// TIA Portal project "TESTV18" (V18) (continued)
REGION Network 13: Bit X12 = Allarme 13
   #_w1 := #IV_CND_ALLX12 AND NOT #VW_Allarms.%X12;
   #TI_T12.TON(IN := #_w1, PT := T#5S);
   IF #_w1 AND #TI_T12.Q THEN
       #VW_Allarms.%X12 := TRUE;   // SR flip-flop
   END_IF;
   IF #IV_RST_ALL THEN #VW_Allarms.%X12 := FALSE; END_IF;
END_REGION

REGION Network 14: Bit X13 = Allarme 14
   #_w1 := #IV_CND_ALLX13 AND NOT #VW_Allarms.%X13;
   #TI_T13.TON(IN := #_w1, PT := T#5S);
   IF #_w1 AND #TI_T13.Q THEN
       #VW_Allarms.%X13 := TRUE;   // SR flip-flop
   END_IF;
   IF #IV_RST_ALL THEN #VW_Allarms.%X13 := FALSE; END_IF;
END_REGION

REGION Network 15: Bit X14 = Allarme 15
   #_w1 := #IV_CND_ALLX14 AND NOT #VW_Allarms.%X14;
   #TI_T14.TON(IN := #_w1, PT := T#5S);
   IF #_w1 AND #TI_T14.Q THEN
       #VW_Allarms.%X14 := TRUE;   // SR flip-flop
   END_IF;
   IF #IV_RST_ALL THEN #VW_Allarms.%X14 := FALSE; END_IF;
END_REGION

REGION Network 16: Bit X15 = Allarme 16
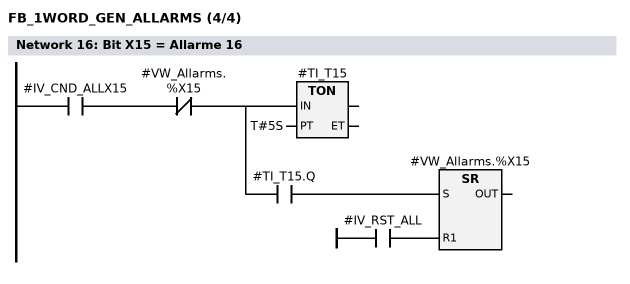
   #_w1 := #IV_CND_ALLX15 AND NOT #VW_Allarms.%X15;
   #TI_T15.TON(IN := #_w1, PT := T#5S);
   IF #_w1 AND #TI_T15.Q THEN
       #VW_Allarms.%X15 := TRUE;   // SR flip-flop
   END_IF;
   IF #IV_RST_ALL THEN #VW_Allarms.%X15 := FALSE; END_IF;
END_REGION
END_FUNCTION_BLOCK

FUNCTION_BLOCK "FB_CYL_DIAGN"   // FB550, LAD
TITLE = FB_CYL_DIAGN
{ S7_Optimized_Access := 'TRUE' }
AUTHOR : C.M.
VERSION : 0.1
// FB per diagnostica cilindro
   VAR_INPUT
      PMI_Limit_Switch_Backward : Bool := FALSE;   // Sensore di posizione cilindro retratto
      PMS_Limit_Switch_Forward : Bool := FALSE;   // Sensore di posizione cilindro esteso
      PST_Home_Position_Backward : Bool := FALSE;   // Posizione HOME indietro
      PST_Home_Position_Forward : Bool := FALSE;   // Posizione HOME avanti
      PST_Latch_In_Backward_Position : Bool := FALSE;   // Interlock in posizione indietro
      PST_Latch_In_Forward_Position : Bool := FALSE;   // Interlock in posizione avanti
      PST_Alarm_Muting : Bool;   // Interlock per sospensione allarmi
      IV_CMD_EV_BCK : Bool;   // Ingresso per conferma attivazione comando cilindro retratto
      IV_CMD_EV_FWD : Bool;   // Ingresso per conferma attivazione comando cilindro esteso
      Station_Info : "Machine_Status_Data";   // Informazioni generali stazione
   END_VAR
   VAR_OUTPUT
      VW_AllarmDIA : Word;   // Variabile WORD per allarmi
   END_VAR
   VAR
      CIN_Auto_Request_Backward : Bool := FALSE;
      CIN_Auto_Request_Forward : Bool := FALSE;
      CIN_Manual_PB_Request_Backward : Bool := FALSE;
      CIN_Manual_PB_Request_Forward : Bool := FALSE;
      CYL_In_Backward_Position : Bool := FALSE;
      CYL_In_Forward_Position : Bool := FALSE;
      CYL_In_Home_Position : Bool := FALSE;
      LOC_SensorBackup_Backward : Bool := FALSE;
      LOC_SensorBackup_Forward : Bool := FALSE;
      LOC_Pulse_1 : Bool;
      LOC_Pulse_2 : Bool;
   END_VAR
   VAR RETAIN
      LOC_DiagnDelay_Backward : Time := T#5s;
      LOC_DiagnDelay_Forward : Time := T#5s;
   END_VAR
   VAR
      LOC_Timer_NotReached_Backward : IEC_TIMER;
      LOC_Timer_NotReached_Forward : IEC_TIMER;
      LOC_Timer_SwitchesContemp : IEC_TIMER;
   END_VAR
   VAR RETAIN
      DIA : "Cylinder_Diagnostic";
   END_VAR
   VAR_TEMP
      No_error : Bool;
   END_VAR
   VAR_TEMP   // added for the SCL form of the ladder/FBD networks
      _w1 : Bool;
   END_VAR
BEGIN

REGION Network 1: *** STATO FINECORSA ***
END_REGION

REGION Network 2: LOGICA - movimento indietro eseguito
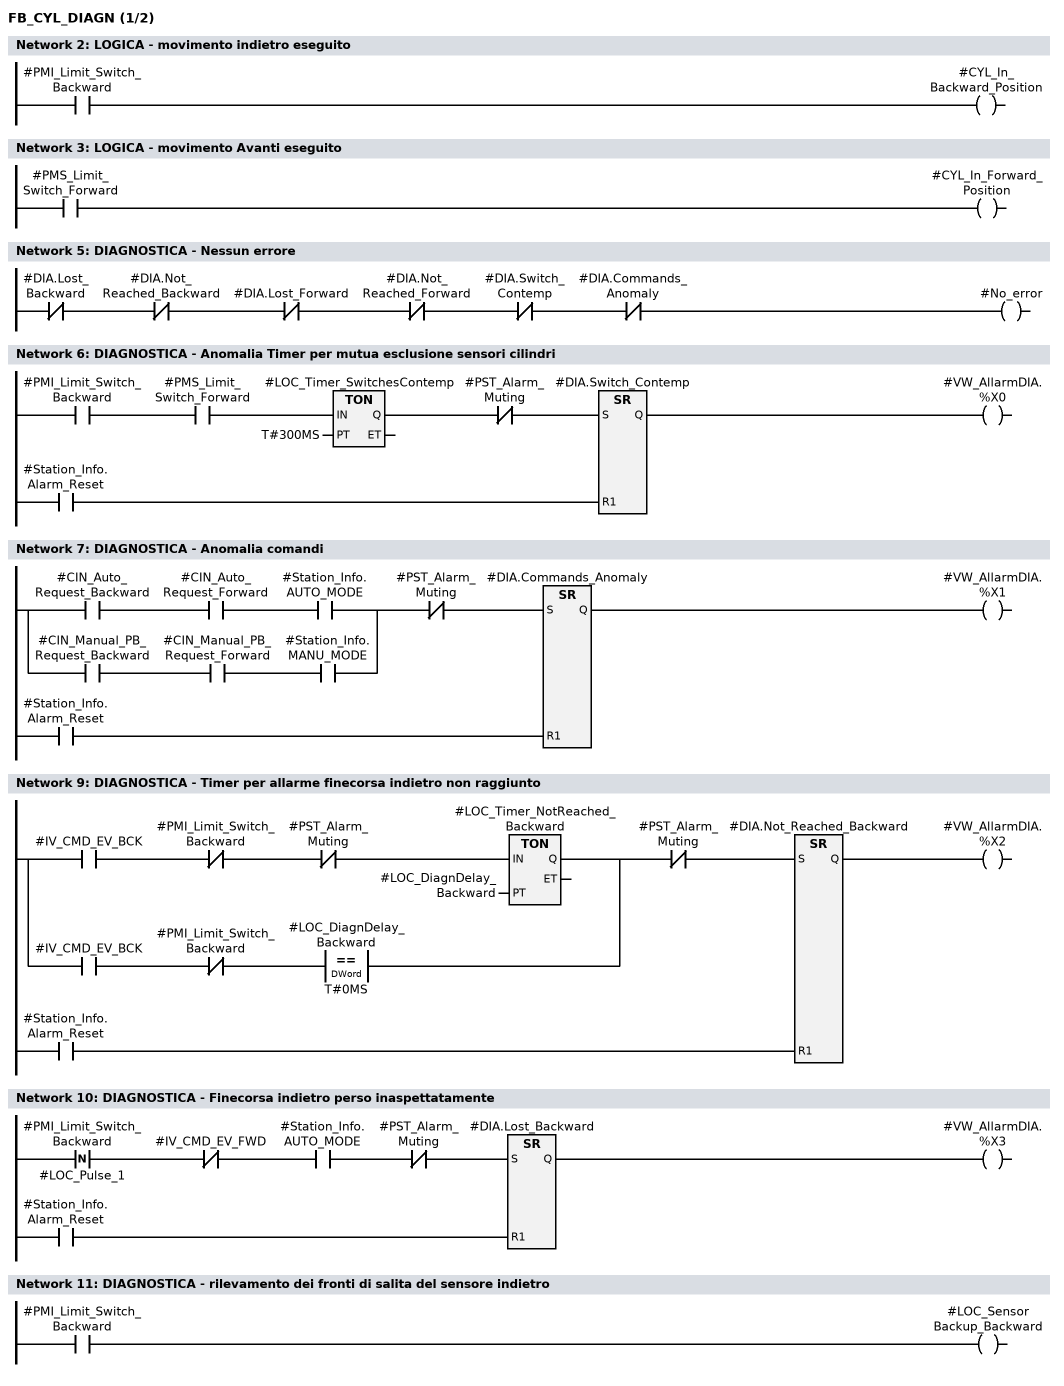
   RUNG wire#powerrail
      Contact( #PMI_Limit_Switch_Backward )
      Coil( #CYL_In_Backward_Position )
   END_RUNG
   // the same network as SCL:
   #CYL_In_Backward_Position := #PMI_Limit_Switch_Backward;
END_REGION

REGION Network 3: LOGICA - movimento Avanti eseguito
   RUNG wire#powerrail
      Contact( #PMS_Limit_Switch_Forward )
      Coil( #CYL_In_Forward_Position )
   END_RUNG
   // the same network as SCL:
   #CYL_In_Forward_Position := #PMS_Limit_Switch_Forward;
END_REGION

REGION Network 4: *** DIAGNOSTICA ***
END_REGION

REGION Network 5: DIAGNOSTICA - Nessun errore
   RUNG wire#powerrail
      I_Contact( #DIA.Lost_Backward )
      I_Contact( #DIA.Not_Reached_Backward )
      I_Contact( #DIA.Lost_Forward )
      I_Contact( #DIA.Not_Reached_Forward )
      I_Contact( #DIA.Switch_Contemp )
      I_Contact( #DIA.Commands_Anomaly )
      Coil( #No_error )
   END_RUNG
   // the same network as SCL:
   #No_error := NOT #DIA.Lost_Backward AND NOT #DIA.Not_Reached_Backward AND NOT #DIA.Lost_Forward AND NOT #DIA.Not_Reached_Forward AND NOT #DIA.Switch_Contemp AND NOT #DIA.Commands_Anomaly;
END_REGION

REGION Network 6: DIAGNOSTICA - Anomalia Timer per mutua esclusione sensori cilindri
   #LOC_Timer_SwitchesContemp.TON(IN := #PMI_Limit_Switch_Backward AND #PMS_Limit_Switch_Forward, PT := T#300MS);
   IF #LOC_Timer_SwitchesContemp.Q AND NOT #PST_Alarm_Muting THEN
       #DIA.Switch_Contemp := TRUE;   // SR flip-flop
   END_IF;
   IF #Station_Info.Alarm_Reset THEN #DIA.Switch_Contemp := FALSE; END_IF;
   #VW_AllarmDIA.%X0 := #DIA.Switch_Contemp;
END_REGION

REGION Network 7: DIAGNOSTICA - Anomalia comandi
   RUNG wire#powerrail
      Contact( #CIN_Auto_Request_Backward )
      Contact( #CIN_Auto_Request_Forward )
      Contact( #Station_Info.AUTO_MODE )
      wire#w1
      I_Contact( #PST_Alarm_Muting )
      S_SR(operand := #DIA.Commands_Anomaly, r1 := wire#w2)
      Coil( #VW_AllarmDIA.%X1 )
   END_RUNG
   RUNG wire#powerrail
      Contact( #CIN_Manual_PB_Request_Backward )
      Contact( #CIN_Manual_PB_Request_Forward )
      Contact( #Station_Info.MANU_MODE )
   END_RUNG wire#w1
   RUNG wire#powerrail
      Contact( #Station_Info.Alarm_Reset )
   END_RUNG wire#w2
   // the same network as SCL:
   IF ((#CIN_Auto_Request_Backward AND #CIN_Auto_Request_Forward AND #Station_Info.AUTO_MODE) OR (#CIN_Manual_PB_Request_Backward AND #CIN_Manual_PB_Request_Forward AND #Station_Info.MANU_MODE)) AND NOT #PST_Alarm_Muting THEN
       #DIA.Commands_Anomaly := TRUE;   // SR flip-flop
   END_IF;
   IF #Station_Info.Alarm_Reset THEN #DIA.Commands_Anomaly := FALSE; END_IF;
   #VW_AllarmDIA.%X1 := #DIA.Commands_Anomaly;
END_REGION

REGION Network 8: *** DIAGNOSTICA SENSORE INDIETRO PMI ***
END_REGION

REGION Network 9: DIAGNOSTICA - Timer per allarme finecorsa indietro non raggiunto
   #LOC_Timer_NotReached_Backward.TON(IN := #IV_CMD_EV_BCK AND NOT #PMI_Limit_Switch_Backward AND NOT #PST_Alarm_Muting,
                           PT := #LOC_DiagnDelay_Backward);
   IF (#LOC_Timer_NotReached_Backward.Q OR (#IV_CMD_EV_BCK AND NOT #PMI_Limit_Switch_Backward AND (#LOC_DiagnDelay_Backward = T#0MS))) AND NOT #PST_Alarm_Muting THEN
       #DIA.Not_Reached_Backward := TRUE;   // SR flip-flop
   END_IF;
   IF #Station_Info.Alarm_Reset THEN #DIA.Not_Reached_Backward := FALSE; END_IF;
   #VW_AllarmDIA.%X2 := #DIA.Not_Reached_Backward;
END_REGION

REGION Network 10: DIAGNOSTICA - Finecorsa indietro perso inaspettatamente
   RUNG wire#powerrail
      N_Contact(operand := #PMI_Limit_Switch_Backward, bit := #LOC_Pulse_1)
      I_Contact( #IV_CMD_EV_FWD )
      Contact( #Station_Info.AUTO_MODE )
      I_Contact( #PST_Alarm_Muting )
      S_SR(operand := #DIA.Lost_Backward, r1 := wire#w1)
      Coil( #VW_AllarmDIA.%X3 )
   END_RUNG
   RUNG wire#powerrail
      Contact( #Station_Info.Alarm_Reset )
   END_RUNG wire#w1
   // the same network as SCL:
   #_w1 := NOT #PMI_Limit_Switch_Backward AND #LOC_Pulse_1;   // falling edge of #PMI_Limit_Switch_Backward
   #LOC_Pulse_1 := #PMI_Limit_Switch_Backward;
   IF #_w1 AND NOT #IV_CMD_EV_FWD AND #Station_Info.AUTO_MODE AND NOT #PST_Alarm_Muting THEN
       #DIA.Lost_Backward := TRUE;   // SR flip-flop
   END_IF;
   IF #Station_Info.Alarm_Reset THEN #DIA.Lost_Backward := FALSE; END_IF;
   #VW_AllarmDIA.%X3 := #DIA.Lost_Backward;
END_REGION

REGION Network 11: DIAGNOSTICA - rilevamento dei fronti di salita del sensore indietro
   RUNG wire#powerrail
      Contact( #PMI_Limit_Switch_Backward )
      Coil( #LOC_SensorBackup_Backward )
   END_RUNG
   // the same network as SCL:
   #LOC_SensorBackup_Backward := #PMI_Limit_Switch_Backward;
END_REGION

REGION Network 12: *** DIAGNOSTICA SENSORE AVANTI PMS ***
END_REGION

REGION Network 13: DIAGNOSTICA - Timer per allarme finecorsa avanti non raggiunto
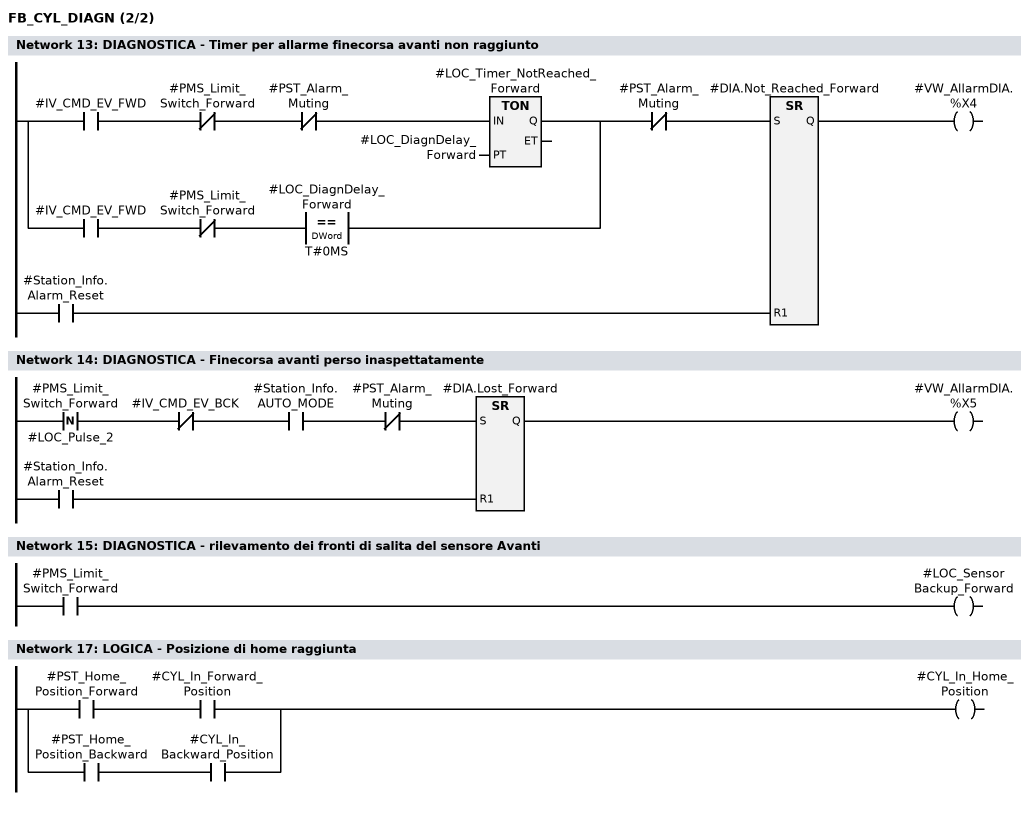
   #LOC_Timer_NotReached_Forward.TON(IN := #IV_CMD_EV_FWD AND NOT #PMS_Limit_Switch_Forward AND NOT #PST_Alarm_Muting,
                           PT := #LOC_DiagnDelay_Forward);
   IF (#LOC_Timer_NotReached_Forward.Q OR (#IV_CMD_EV_FWD AND NOT #PMS_Limit_Switch_Forward AND (#LOC_DiagnDelay_Forward = T#0MS))) AND NOT #PST_Alarm_Muting THEN
       #DIA.Not_Reached_Forward := TRUE;   // SR flip-flop
   END_IF;
   IF #Station_Info.Alarm_Reset THEN #DIA.Not_Reached_Forward := FALSE; END_IF;
   #VW_AllarmDIA.%X4 := #DIA.Not_Reached_Forward;
END_REGION

REGION Network 14: DIAGNOSTICA - Finecorsa avanti perso inaspettatamente
   RUNG wire#powerrail
      N_Contact(operand := #PMS_Limit_Switch_Forward, bit := #LOC_Pulse_2)
      I_Contact( #IV_CMD_EV_BCK )
      Contact( #Station_Info.AUTO_MODE )
      I_Contact( #PST_Alarm_Muting )
      S_SR(operand := #DIA.Lost_Forward, r1 := wire#w1)
      Coil( #VW_AllarmDIA.%X5 )
   END_RUNG
   RUNG wire#powerrail
      Contact( #Station_Info.Alarm_Reset )
   END_RUNG wire#w1
   // the same network as SCL:
   #_w1 := NOT #PMS_Limit_Switch_Forward AND #LOC_Pulse_2;   // falling edge of #PMS_Limit_Switch_Forward
   #LOC_Pulse_2 := #PMS_Limit_Switch_Forward;
   IF #_w1 AND NOT #IV_CMD_EV_BCK AND #Station_Info.AUTO_MODE AND NOT #PST_Alarm_Muting THEN
       #DIA.Lost_Forward := TRUE;   // SR flip-flop
   END_IF;
   IF #Station_Info.Alarm_Reset THEN #DIA.Lost_Forward := FALSE; END_IF;
   #VW_AllarmDIA.%X5 := #DIA.Lost_Forward;
END_REGION

REGION Network 15: DIAGNOSTICA - rilevamento dei fronti di salita del sensore Avanti
   RUNG wire#powerrail
      Contact( #PMS_Limit_Switch_Forward )
      Coil( #LOC_SensorBackup_Forward )
   END_RUNG
   // the same network as SCL:
   #LOC_SensorBackup_Forward := #PMS_Limit_Switch_Forward;
END_REGION

REGION Network 16: *** SEGMENTI DI LOGICA AUSILIARI ***
END_REGION

REGION Network 17: LOGICA - Posizione di home raggiunta
   RUNG wire#powerrail
      Contact( #PST_Home_Position_Forward )
      Contact( #CYL_In_Forward_Position )
      wire#w1
      Coil( #CYL_In_Home_Position )
   END_RUNG
   RUNG wire#powerrail
      Contact( #PST_Home_Position_Backward )
      Contact( #CYL_In_Backward_Position )
   END_RUNG wire#w1
   // the same network as SCL:
   #CYL_In_Home_Position := (#PST_Home_Position_Forward AND #CYL_In_Forward_Position) OR (#PST_Home_Position_Backward AND #CYL_In_Backward_Position);
END_REGION
END_FUNCTION_BLOCK

// folder: LGF/1 Date and timer operations

FUNCTION "LGF_GetCalendarDay" : DInt   // FC10028, SCL
TITLE = LGF_GetCalendarDay
{ S7_Optimized_Access := 'TRUE' }
AUTHOR : Siemens_Digital_Industry
FAMILY : LGF
NAME : LGF_GetCalendarDay
// This function uses the specified date to calculate the number of days that have passed since the beginning of the year (1st January).
// 
// The function is used in the functions “LGF_GetCalendarWeek_ISO” and “LGF_GetCalendarWeek_US”.
// Diese Funktion berechnet aus dem vorgegebenen Datum die Anzahl der Tage, die seit dem Anfang des Jahres vergangen sind (1. Januar).
// 
// Die Funktion wird in den Funktionen "LGF_GetCalendarWeek_ISO" und "LGF_GetCalendarWeek_US" verwendet.
   VAR_INPUT
      "date" : DTL;   // Date for the calculation of the calendar days since 1 January. / Datum für die Berechnung der vergangenen Kalendertagen seit dem 01. Januar
   END_VAR
   VAR_OUTPUT
      error : Bool;   // FALSE: No error / TRUE: An error occurred during the execution of the FB / FALSE: Kein Fehler / TRUE: Während der Ausführung des FB ist ein Fehler aufgetreten
      status : Word;   // 16#0000-16#7FFF: Status of the FB / 16#8000-16#FFFF: Error identification (see following Table) / 16#0000-16#7FFF: Status des FB / 16#8000-16#FFFF: Fehleridentifikation (siehe folgende Tabelle)
   END_VAR
   VAR_TEMP
      tempDaysPassed : DInt;   // Temp tag for the number of days past / Temp Variable für die Anzahl der vergangenen Tage
      tempDate : DTL;   // Temp variable to store date for calculations / Temp Variable um Datum für Berechung zwischen zu speichern
   END_VAR
   // Ret_Val : Days past since January 1st. / Vergangene Tage seit 1. Januar.
   VAR CONSTANT
      FIRST_DAY : USInt := 1;   // 1st of a month / 1. Tag eines Monats
      LAST_DAY : USInt := 31;   // 31st of a month / 31. Tag eines Monats
      JANUARY : USInt := 1;   // Month number for January / Monatsnumer Januar
      DECEMBER : USInt := 12;   // Month number for December / Monatsnummer Dezember
      TIME_ZERO_FORCE_UPDATE : Time := t#0d;   // By adding zero an update of DTL Tag is forced and auto checks are applied / Durch die Addition von "0" wird ein Update üder den Zeitstemple erstellt und ebenfalls auf gültigkeit geprüft.
      ONE_DAY : DInt := 1;   // One single day for incrementing / Ein Tag für inkrementierungen
      STATUS_NO_ERROR : Word := 16#0000;   // Status: no error occurred / Status: kein Fehler aufgetreten
      ERR_LIM_DATE : Word := 16#8201;   // Date out of the range, has to be greater than <1970-01-01 ; 2262-04-11> / Datum ausserhalb des gültigen Bereiches, es muss nach dem <1970-01-01 ; 2262-04-11> liegen
   END_VAR
BEGIN
   REGION BLOCK INFO HEADER
     //===============================================================================
     // SIEMENS AG / (c)Copyright 2019
     //-------------------------------------------------------------------------------
     // Title:            LGF_GetCalendarDay
     // Comment/Function: This function calculates for a date the passed days since 1st January.
     // Library/Family:   LGF(Library General Functions)
     // Author:           Siemens Digital Industry Support
     // Tested with:      S7-PLCSIM Advanced V2.0 SP1
     // Engineering:      TIA Portal V15.1
     // Restrictions:     ENO disabled - error handling done with error and status
     // Requirements:     PLC (S7-1200 / S7-1500)
     //-------------------------------------------------------------------------------
     // Change log table:
     // Version  | Date       | Expert in charge       | Changes applied
     //----------|------------|------------------------|------------------------------
     // 01.00.00 16.07.2019  Simatic Systems Support
     //                      First release
     //                      ENO used for internal error handling, interface has error and status
     //                      temp tag naming, insert constant
     // 03.00.00 23.04.2020  Simatic Systems Support
     //                      Set version to V3.0.0, harmonize the version of the whole library
     // 03.00.01 19.01.2020  Simatic Systems Support
     //                      Insert documentation
     //=============================================================================
   END_REGION BLOCK INFO HEADER

   REGION INITIALISATION
     #tempDate := #date;
     #tempDaysPassed := 0;
   END_REGION

   REGION COUNT DAYS
     // Check #date
     // adding zero forces the PLC to update the tag and eno check
     #tempDate := #tempDate + #TIME_ZERO_FORCE_UPDATE;
     IF ENO = FALSE THEN
       #error := TRUE;
       #status := #ERR_LIM_DATE;
       #LGF_GetCalendarDay := #tempDaysPassed;
       RETURN;
     END_IF;

     // Weekday of 1st January in the current year
     #tempDate.MONTH := #JANUARY;
     #tempDate.DAY := #FIRST_DAY;
     // adding zero forces the PLC to update the tag
     // in this case especially the weekday
     #tempDate := #tempDate + #TIME_ZERO_FORCE_UPDATE;

     // Days passed in the year since 1st January, "date" included
     #tempDaysPassed := DATE_TO_DINT(DTL_TO_DATE(#date)) - DATE_TO_DINT(DTL_TO_DATE(#tempDate)) + #ONE_DAY;
   END_REGION

   REGION OUTPUTS
     #error := FALSE;
     #status := #STATUS_NO_ERROR;
     #LGF_GetCalendarDay := #tempDaysPassed;

     // ENO is not used, forced to TRUE
     ENO := TRUE;
   END_REGION
END_FUNCTION

// folder: LGF/4 Math operations

FUNCTION "LGF_CalcDistance_2D" : LReal   // FC10020, SCL
TITLE = LGF_CalcDistance_2D
{ S7_Optimized_Access := 'TRUE' }
AUTHOR : Siemens_Digital_Industries
FAMILY : LGF
NAME : LGF_CalcDistance_2D
// The function calculates the distance between two points in the plane. / Die Funktion berechnet den Abstand zwischen zwei Punkten in der Ebene.
   VAR_INPUT
      x1 : LReal;   // X coordinate point 1 / X Koordinate Punkt 1
      y1 : LReal;   // Y coordinate point 1 / Y Koordinate Punkt 1
      x2 : LReal;   // X coordinate point 2 / X Koordinate Punkt 2
      y2 : LReal;   // Y coordinate point 2 / Y Koordinate Punkt 2
   END_VAR
   // Ret_Val : Calculated distance between the Points / Berechnete Distanz zwischen den Punkten
BEGIN
   REGION Block info header
     //=============================================================================
     // Siemens AG / (c)Copyright 2017
     //-----------------------------------------------------------------------------
     // Title:            LGF_CalcDistance_2D
     // Comment/Function: Calculates the distance between two points in 2D space
     // Library/Family:   LGF(Library General Functions)
     // Author:           Siemens Digital Industry Support
     // Tested with:      S7-PLCSIM Advanced V2.0 SP1
     // Engineering:      TIA Portal V15 Update 2
     // Restrictions:     ENO disabled - ENO mechanism is not used
     // Requirements:     PLC (S7-1200 / S7-1500)
     //-------------------------------------------------------------------------------
     // Change log table:
     // Version  | Date       | Expert in charge       | Changes applied
     //----------|------------|------------------------|------------------------------
     // 01.00.00 06.07.2018  Siemens Industry Online Support
     //                      First released version
     // 01.00.01 17.08.2018  Siemens Industry Online Support
     //                      Upgrade: TIA V15 Update 2
     // 01.00.02 23.11.2018  Siemens Industry Online Support
     //                      Upgrade: TIA V15.1
     // 01.02.00 04.10.2019  Simatic Systems Support
     //                      renamed from "Distance" to "CalcDistance_2D"
     //                      Data type changed to LREAL
     //                      Data type changed to LREAL
     // 03.00.00 23.04.2020  Simatic Systems Support
     //                      Set version to V3.0.0, harmonize the version of the whole library
     // 03.00.01 12.11.2020  Simatic Systems Support
     //                      Insert documentation
     //=============================================================================
   END_REGION Block info header

   REGION DESCRIPTION
     (/*The block calculates the distance between two points in a Cartesian coordinate system. The distance is calculated with the following formula:

   $$
    result = \sqrt[2]{(x_2-x_1)^2+(y_2-y_1)^2}
   $$

   ------

   Figure: Graphical representation

   ![LGF_CalcDistance_2D - Principle of operation](LGF_CalcDistance_2D.PNG "LGF_CalcDistance_2D - Principle of operation")
   Der Baustein berechnet den Abstand zwischen zwei Punkten in einem kartesischen Koordinatensystem. Der Abstand wird mit nachfolgender Formel berechnet:

   $$
    result = \sqrt[2]{(x_2-x_1)^2+(y_2-y_1)^2}
   $$

   ------

   Abbildung: Graphische Darstellung

   ![LGF_CalcDistance_2D - Funktionsweise](LGF_CalcDistance_2D.PNG "LGF_CalcDistance_2D - Funktionsweise")*/)
   END_REGION DESCRIPTION

   REGION Program
     // Calculating the distance
     #LGF_CalcDistance_2D := SQRT(SQR(#x2 - #x1) + SQR(#y2 - #y1));
     // ENO mechanism is not used
     ENO := TRUE;
   END_REGION
END_FUNCTION

// folder: LGF/6 Converter operations

FUNCTION "LGF_BinaryToGray" : DWord   // FC10021, SCL
TITLE = LGF_BinaryToGray
{ S7_Optimized_Access := 'TRUE' }
AUTHOR : Siemens_Digital_Industry
FAMILY : LGF
NAME : LGF_BinaryToGray
// This function converts a binary coded value into a Gray-coded value. / Diese Funktion wandelt einen binär codierten Wert in einen Gray codierten Wert um.
   VAR_INPUT
      variableBinary : DWord;   // Binary coded value to convert to Gray code / Binär codierter Wert der zu Gray-Code umgerechnet wird
   END_VAR
   // Ret_Val : Gray-coded value / Gray codierter Wert
   VAR CONSTANT
      BIT_SHIFT_1 : USInt := 1;   // The number (1) of bit positions by which the specified value should be shifted.
   END_VAR
BEGIN
   REGION BLOCK INFO HEADER
     //===============================================================================
     // SIEMENS AG / (c)Copyright 2017
     //-------------------------------------------------------------------------------
     // Title:            LGF_BinaryToGray
     // Comment/Function: This function converts a binary value to a gray coded value
     // Library/Family:   LGF(Library General Functions)
     // Author:           Siemens Digital Industry Support
     // Tested with:      CPU1212C DC/DC/DC FW:V4.2
     // Engineering:      TIA Portal V14 Update 1
     // Restrictions:     ENO disabled - no error handling needed
     // Requirements:     PLC (S7-1200 / S7-1500)
     //-------------------------------------------------------------------------------
     // Change log table:
     // Version  | Date       | Expert in charge       | Changes applied
     //----------|------------|------------------------|------------------------------
     // 01.00.00 | 19.08.2015 | Siemens Industry Online Support
     //                         First released version
     // 01.00.01 | 28.10.2015 | Siemens Industry Online Support
     //                         Name changed
     // 01.00.02 | 02.01.2017 | Siemens Industry Online Support
     //                         Upgrade: TIA Portal V14 Update 1
     // 01.00.03 | 17.08.2018 | Siemens Industry Online Support
     //                         Upgrade: TIA V15 Update 2
     // 01.00.04 | 23.11.2018 | Siemens Industry Online Support
     //                         Upgrade: TIA V15.1
     // 01.00.05 | 11.06.2019 | Simatic Systems Support
     //                         Standard header and block parameters update
     //                         Add ENO handling
     // 03.00.00 | 23.04.2020 | Simatic Systems Support | Set version to V3.0.0
     //                         Harmonize the version of the whole library
     // 03.00.01 | 23.02.2021 | Simatic Systems Support
     //                         Insert documentation
     //===============================================================================
   END_REGION Block info header

   REGION OUTPUTS
     #LGF_BinaryToGray := #variableBinary XOR SHR(IN := #variableBinary, N := #BIT_SHIFT_1);

     // no error handling needed
     ENO := TRUE;
   END_REGION
END_FUNCTION

// folder: LGF/6 Converter operations/Binary types - Split/Merge

FUNCTION "LGF_MergeBitsToByte" : Byte   // FC10060, SCL
TITLE = LGF_MergeBitsToByte
{ S7_Optimized_Access := 'TRUE' }
AUTHOR : Siemens_Digital_Industry
FAMILY : LGF
NAME : LGF_MergeBitsToByte
// This function merge 8 Bits / 8 Boolean variables into one Byte variable. / Diese Funktion führt 8 Bit / 8 Boolsche Variablen in einer Byte Variable zusammen.
   VAR_INPUT
      bit7 : Bool;   // Input Bit 7 - MSB
      bit6 : Bool;   // Input Bit 6
      bit5 : Bool;   // Input Bit 5
      bit4 : Bool;   // Input Bit 4
      bit3 : Bool;   // Input Bit 3
      bit2 : Bool;   // Input Bit 2
      bit1 : Bool;   // Input Bit 1
      bit0 : Bool;   // Input Bit 0 - LSB
   END_VAR
   VAR_TEMP
      tempByte : Byte;   // Temp memory to merge Bits into a Byte / Temp speicher zum zusammenführen der Bits zu einem Byte
   END_VAR
   // Ret_Val : Composite Bit sequence stored as Byte variable / Zusammengefügte Bitfolge, gespeichert in einer Byte Variable
BEGIN
   REGION BLOCK INFO HEADER
     //===============================================================================
     // SIEMENS AG / (c)Copyright 2018
     //-------------------------------------------------------------------------------
     // Title:            LGF_MergeBitsToByte
     // Comment/Function: This function merge 8 Bits / 8 Boolean variables into one Byte variable.
     // Library/Family:   LGF (Library General Functions)
     // Author:           Siemens Digital Industry Support
     // Tested with:      S7-PLCSIM Advanced V2.0 SP1
     // Engineering:      TIA Portal V14 / V14SP1
     // Restrictions:     ENO disabled - no error handling, no failure possible.
     // Requirements:     PLC (S7-1200 / S7-1500)
     //-------------------------------------------------------------------------------
     // Change log table:
     // Version  | Date       | Expert in charge       | Changes applied
     //----------|------------|------------------------|------------------------------
     // 01.00.00 | 20.06.2019 | Simatic Systems Support
     //                         First release
     // 03.00.00 | 23.04.2020 | Simatic Systems Support | Set version to V3.0.0
     //                         harmonize the version of the whole library
     // 03.00.01 | 22.02.2021 | Simatic Systems Support
     //                         Insert documentation
     //=============================================================================
   END_REGION

   REGION MERGE
     // set the bits by slice access
     #tempByte.%X7 := #bit7;
     #tempByte.%X6 := #bit6;
     #tempByte.%X5 := #bit5;
     #tempByte.%X4 := #bit4;
     #tempByte.%X3 := #bit3;
     #tempByte.%X2 := #bit2;
     #tempByte.%X1 := #bit1;
     #tempByte.%X0 := #bit0;
   END_REGION

   REGION OUTPUT
     #LGF_MergeBitsToByte := #tempByte;
     // no error handling needed
     ENO := TRUE;
   END_REGION
END_FUNCTION

FUNCTION "LGF_SplitByteToBits" : Void   // FC10063, SCL
TITLE = LGF_SplitByteToBits
{ S7_Optimized_Access := 'TRUE' }
AUTHOR : Siemens_Digital_Industry
FAMILY : LGF
NAME : LGF_SplitByteToBits
// This function splits a Byte variable into 8 Boolean / 8 Bit variables. / Diese Funktion zerlegt eine Byte Variable in 8 Bool / 8 Bit Variablen.
   VAR_INPUT
      "byte" : Byte;   // Bit sequence to be split / Bitfolge die zerlegt wird
   END_VAR
   VAR_OUTPUT
      bit7 : Bool;   // Output Bit 7 - MSB
      bit6 : Bool;   // Output Bit 6
      bit5 : Bool;   // Output Bit 5
      bit4 : Bool;   // Output Bit 4
      bit3 : Bool;   // Output Bit 3
      bit2 : Bool;   // Output Bit 2
      bit1 : Bool;   // Output Bit 1
      bit0 : Bool;   // Output Bit 0 - LSB
   END_VAR
BEGIN
   REGION BLOCK INFO HEADER
     //===============================================================================
     // SIEMENS AG / (c)Copyright 2018
     //-------------------------------------------------------------------------------
     // Title:            LGF_SplitByteToBits
     // Comment/Function: This function splits a Byte variable into 8 Boolean / 8 Bit variables
     // Library/Family:   LGF (Library General Functions)
     // Author:           Siemens Digital Industry Support
     // Tested with:      S7-PLCSIM Advanced V2.0 SP1
     // Engineering:      TIA Portal V14 / V14SP1
     // Restrictions:     ENO disabled - no error handling, no failure possible.
     // Requirements:     PLC (S7-1200 / S7-1500)
     //-------------------------------------------------------------------------------
     // Change log table:
     // Version  | Date       | Expert in charge       | Changes applied
     //----------|------------|------------------------|------------------------------
     // 01.00.00 | 20.06.2019 | Simatic Systems Support
     //                         First release
     // 03.00.00 | 23.04.2020 | Simatic Systems Support | Set version to V3.0.0
     //                         harmonize the version of the whole library
     // 03.00.01 | 22.02.2021 | Simatic Systems Support
     //                         Insert documentation
     //=============================================================================
   END_REGION

   REGION OUTPUT
     // get the bits by slice access
     #bit7 := #byte.%X7;
     #bit6 := #byte.%X6;
     #bit5 := #byte.%X5;
     #bit4 := #byte.%X4;
     #bit3 := #byte.%X3;
     #bit2 := #byte.%X2;
     #bit1 := #byte.%X1;
     #bit0 := #byte.%X0;
     // no error handling needed
     ENO := TRUE;
   END_REGION
END_FUNCTION

// folder: MTA/Vari

FUNCTION_BLOCK "ALM_VALVE_CFG1"   // FB2, LAD
TITLE = FB gestione allarmi elettrov. con cilindro pneum.
{ S7_Optimized_Access := 'TRUE' }
AUTHOR : Cecini_M
VERSION : 0.1
// ROUTINE DI GESTIONE ALLARMI ELETTROVALVOLA COMBINATA CON CILINDRO PNEUMATICO.
//  - Usare ingressi CMD1 e CMD2 per bistabile. Usare negazione di CMD1 su CMD2 per monost.
//  - Ingressi di timeout in S 0.0 (convertiti all'interno dell'FB)
//  - 2 CMD Valvola + 2 Sensori posizione SM
//  - Allarme mancanza sensore su CMD1
//  - Allarme mancanza sensore su CMD2
//  - Allarme mutua eslusione entrambi SM
   VAR_INPUT
      IV_YV_CMD1 : Bool;   // Ingresso comando direzione 1
      IV_YV_CMD2 : Bool;   // Ingresso comando direzione 2
      IV_FBK_CMD1 : Bool;   // Ingresso sensore SM comando direzione 1
      IV_FBK_CMD2 : Bool;   // Ingresso sensore SM comando direzione 1
   END_VAR
   VAR_OUTPUT
      Vb_ALM1 : Bool;
      Vb_ALM2 : Bool;
      Vb_ALM3 : Bool;
   END_VAR
   VAR_IN_OUT
      IV_ACK_ALM1 : Bool;   // Ingresso ACK riconoscimento ALM1
      IV_ACK_ALM2 : Bool;   // Ingresso ACK riconoscimento ALM2
      IV_ACK_ALM3 : Bool;   // Ingresso ACK riconoscimento ALM3
      TI_ToutALM1 : UInt;   // Timeout allarme1
      TI_ToutALM2 : UInt;   // Timeout allarme2
      TI_ToutALM3 : UInt;   // Timeout allarme3
   END_VAR
   VAR
      TI_T1 : IEC_TIMER;   // Timer ALM1
      TI_T2 : IEC_TIMER;   // Timer ALM1
      TI_T3 : IEC_TIMER;   // Timer ALM1
      ME_ALM1 : Bool;   // Memoria allarme 1 SM CMD1
      ME_ALM2 : Bool;   // Memoria allarme 2 SM CMD2
      ME_ALM3 : Bool;   // Memoria allarme 3 mutua esclusione sensori SM
      VA_SetP_TIALM1 : DInt;   // Valore di SETPOINT per timer ALM1
      VA_SetP_TIALM2 : DInt;   // Valore di SETPOINT per timer ALM2
      VA_SetP_TIALM3 : DInt;   // Valore di SETPOINT per timer ALM3
   END_VAR
   VAR_TEMP
      VA_AppRis1 : UInt;   // Variabile appoggio risultato intermedio 1
      VA_AppRis2 : UInt;   // Variabile appoggio risultato intermedio 2
      VA_AppRis3 : UInt;   // Variabile appoggio risultato intermedio 3
   END_VAR
   VAR_TEMP   // added for the SCL form of the ladder/FBD networks
      _w1 : Bool;
      _w2 : Bool;
   END_VAR
BEGIN

REGION Network 1: Conversione ingressi TIMEOUT in S a MS per IEC TIMER
   // Valori d'ingresso espressi in S 0.0
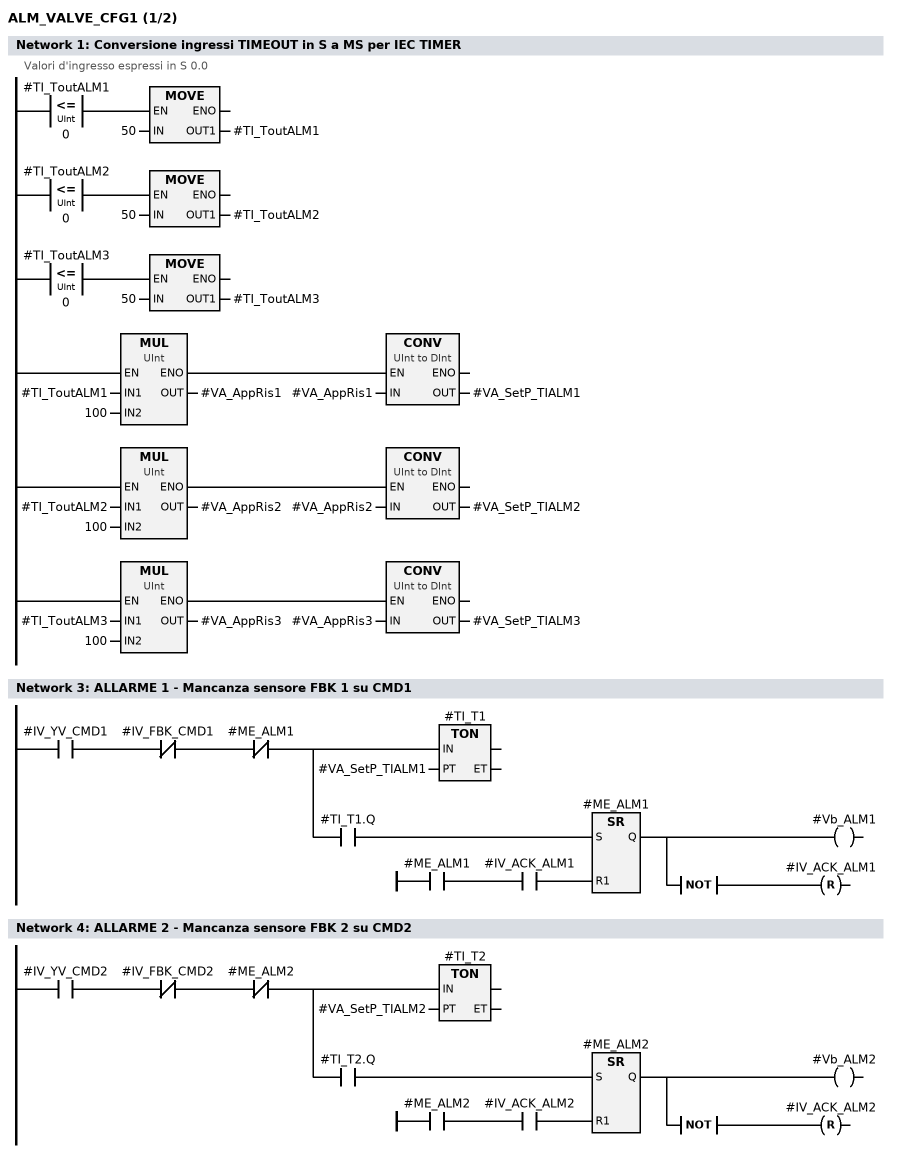
   RUNG wire#powerrail
      { S7_Templates := "SrcType := UInt" } LE_Contact(in1 := #TI_ToutALM1, in2 := 0)
      Move(in := 50, out1 => #TI_ToutALM1)
   END_RUNG
   RUNG wire#powerrail
      { S7_Templates := "SrcType := UInt" } LE_Contact(in1 := #TI_ToutALM2, in2 := 0)
      Move(in := 50, out1 => #TI_ToutALM2)
   END_RUNG
   RUNG wire#powerrail
      { S7_Templates := "SrcType := UInt" } LE_Contact(in1 := #TI_ToutALM3, in2 := 0)
      Move(in := 50, out1 => #TI_ToutALM3)
   END_RUNG
   RUNG wire#powerrail
      { S7_Templates := "SrcType := UInt" } Mul(in1 := #TI_ToutALM1, in2 := 100, out => #VA_AppRis1)
      { S7_Templates := "[SrcType := UInt, DestType := DInt]" } Convert(in := #VA_AppRis1, out => #VA_SetP_TIALM1)
   END_RUNG
   RUNG wire#powerrail
      { S7_Templates := "SrcType := UInt" } Mul(in1 := #TI_ToutALM2, in2 := 100, out => #VA_AppRis2)
      { S7_Templates := "[SrcType := UInt, DestType := DInt]" } Convert(in := #VA_AppRis2, out => #VA_SetP_TIALM2)
   END_RUNG
   RUNG wire#powerrail
      { S7_Templates := "SrcType := UInt" } Mul(in1 := #TI_ToutALM3, in2 := 100, out => #VA_AppRis3)
      { S7_Templates := "[SrcType := UInt, DestType := DInt]" } Convert(in := #VA_AppRis3, out => #VA_SetP_TIALM3)
   END_RUNG
   // the same network as SCL:
   IF #TI_ToutALM1 <= 0 THEN #TI_ToutALM1 := 50; END_IF;
   IF #TI_ToutALM2 <= 0 THEN #TI_ToutALM2 := 50; END_IF;
   IF #TI_ToutALM3 <= 0 THEN #TI_ToutALM3 := 50; END_IF;
   #VA_AppRis1 := #TI_ToutALM1 * 100;
   #VA_SetP_TIALM1 := UINT_TO_DINT(#VA_AppRis1);
   #VA_AppRis2 := #TI_ToutALM2 * 100;
   #VA_SetP_TIALM2 := UINT_TO_DINT(#VA_AppRis2);
   #VA_AppRis3 := #TI_ToutALM3 * 100;
   #VA_SetP_TIALM3 := UINT_TO_DINT(#VA_AppRis3);
END_REGION

REGION Network 2: *** ALLARMI ***
END_REGION

REGION Network 3: ALLARME 1 - Mancanza sensore FBK 1 su CMD1
   #_w1 := #IV_YV_CMD1 AND NOT #IV_FBK_CMD1 AND NOT #ME_ALM1;
   #TI_T1.TON(IN := #_w1, PT := #VA_SetP_TIALM1);
   #_w2 := #ME_ALM1 AND #IV_ACK_ALM1;
   IF #_w1 AND #TI_T1.Q THEN
       #ME_ALM1 := TRUE;   // SR flip-flop
   END_IF;
   IF #_w2 THEN #ME_ALM1 := FALSE; END_IF;
   #Vb_ALM1 := #ME_ALM1;
   IF NOT #ME_ALM1 THEN #IV_ACK_ALM1 := FALSE; END_IF;
END_REGION

REGION Network 4: ALLARME 2 - Mancanza sensore FBK 2 su CMD2
   #_w1 := #IV_YV_CMD2 AND NOT #IV_FBK_CMD2 AND NOT #ME_ALM2;
   #TI_T2.TON(IN := #_w1, PT := #VA_SetP_TIALM2);
   #_w2 := #ME_ALM2 AND #IV_ACK_ALM2;
   IF #_w1 AND #TI_T2.Q THEN
       #ME_ALM2 := TRUE;   // SR flip-flop
   END_IF;
   IF #_w2 THEN #ME_ALM2 := FALSE; END_IF;
   #Vb_ALM2 := #ME_ALM2;
   IF NOT #ME_ALM2 THEN #IV_ACK_ALM2 := FALSE; END_IF;
END_REGION

REGION Network 5: ALLARME 3 - Errore di mutua esclusione FBK. Presenza contemporanea dei due sensori
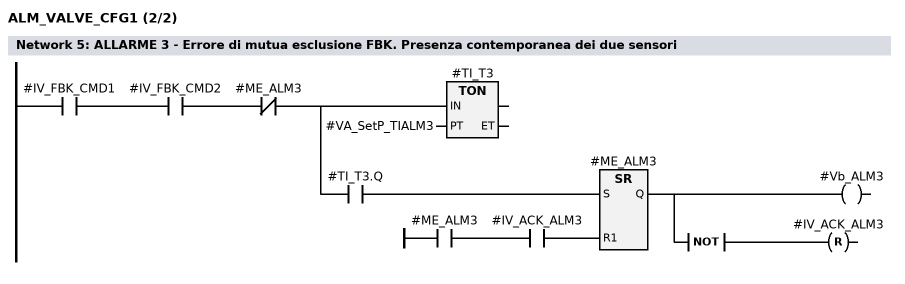
   #_w1 := #IV_FBK_CMD1 AND #IV_FBK_CMD2 AND NOT #ME_ALM3;
   #TI_T3.TON(IN := #_w1, PT := #VA_SetP_TIALM3);
   #_w2 := #ME_ALM3 AND #IV_ACK_ALM3;
   IF #_w1 AND #TI_T3.Q THEN
       #ME_ALM3 := TRUE;   // SR flip-flop
   END_IF;
   IF #_w2 THEN #ME_ALM3 := FALSE; END_IF;
   #Vb_ALM3 := #ME_ALM3;
   IF NOT #ME_ALM3 THEN #IV_ACK_ALM3 := FALSE; END_IF;
END_REGION
END_FUNCTION_BLOCK

// ===== library: CodeBlockByCopyVersionObject "None" =====

// ===== library: CodeBlockByCopyVersionObject "None" =====

// ===== library: CodeBlockByCopyVersionObject "None" =====

// ===== library: CodeBlockByCopyVersionObject "None" =====

// ===== library: CodeBlockByCopyVersionObject "None" =====

// ===== library: CodeBlockByCopyVersionObject "None" =====

// ===== library: CodeBlockByCopyVersionObject "None" =====

